ScreenModuleEditorView "Connection_Parameters_Control" 600x270
   TextField "id_label" at 0,55 size 300x50; Text 'ID'
      Visibility <- "interface.id_label_visible"
      Appearance <- "interface.id_label_animate"
   IOField "id_entry" at 300,55 size 300x50; FormatPattern ??????
      on OnFinishInput: SetBit("interface.id_entry_input_finished")
      on Deactivate: ResetBit("interface.id_entry_active")
      on Activate: SetBit("interface.id_entry_active")
      Appearance <- "interface.id_entry_animate"
      Visibility <- "interface.id_entry_visible"
      ObjectEnable <- "interface.id_entry_enable"
      ProcessValue <- "interface.id_entry_value"
   Button "back" at 0,220 size 600x50; TextOff 'BACK'
      on Press: function_b14e0dd5("interface.back_actuate", 0)
      Appearance <- "interface.back_animate"
      Visibility <- "interface.back_visible"
      ObjectEnable <- "interface.back_enable"
   TextField "ip_address_label" at 0,110 size 300x50; Text 'IP ADDRESS'
      Visibility <- "interface.ip_address_label_visible"
      Appearance <- "interface.ip_address_label_animate"
   IOField "ip_address_entry" at 300,110 size 300x50; FormatPattern ???????????????
      on OnFinishInput: SetBit("interface.ip_address_entry_input_finished")
      on Deactivate: ResetBit("interface.ip_address_entry_active")
      on Activate: SetBit("interface.ip_address_entry_active")
      Appearance <- "interface.ip_address_entry_animate"
      Visibility <- "interface.ip_address_entry_visible"
      ObjectEnable <- "interface.ip_address_entry_enable"
      ProcessValue <- "interface.ip_address_entry_value"
   TextField "port_label" at 0,165 size 300x50; Text 'PORT'
      Visibility <- "interface.port_label_visible"
      Appearance <- "interface.port_label_animate"
   IOField "port_entry" at 300,165 size 300x50; FormatPattern ??????
      on OnFinishInput: SetBit("interface.port_entry_input_finished")
      on Deactivate: ResetBit("interface.port_entry_active")
      on Activate: SetBit("interface.port_entry_active")
      Appearance <- "interface.port_entry_animate"
      Visibility <- "interface.port_entry_visible"
      ObjectEnable <- "interface.port_entry_enable"
      ProcessValue <- "interface.port_entry_value"
   IOField "header" at 0,0 size 600x50; FormatPattern ?????????????????????????
      Appearance <- "interface.header_animate"
      Visibility <- "interface.header_visible"
      ProcessValue <- "interface.header_value"
*)